REGION Network 68: Alarm - Under Range
   RUNG wire#powerrail
      Contact( #Timers.UR_HLD.Q )
      S_SR(operand := #HMI.Alarm.Alarms.%X7, r1 := wire#w1)
   END_RUNG
   RUNG wire#powerrail
      I_Contact( #Timers.UR_HLD.Q )
      { S7_Templates := "SrcType := Real"; S7_GenerateENO := "TRUE" } Add(in1 := #Admin.SCL.UR, in2 := #Retain.HMI.Config.SP.HYS.UR, out => #Admin.HYS.UR)
      { S7_Templates := "SrcType := Real" } GE_Contact(in1 := #RAIVR_1_1, in2 := #Admin.HYS.UR)
   END_RUNG wire#w1
   RUNG wire#powerrail
      I_Contact( #Retain.HMI.Config.Alarms.%X7 )
   END_RUNG wire#w1
   // the same network as SCL:
   // ENO of a box is taken as its EN; it also drops when the box reports an error
   IF NOT #Timers.UR_HLD.Q THEN #Admin.HYS.UR := #Admin.SCL.UR + #Retain.HMI.Config.SP.HYS.UR; END_IF;
   IF #Timers.UR_HLD.Q THEN
       #HMI.Alarm.Alarms.%X7 := TRUE;   // SR flip-flop
   END_IF;
   IF (NOT #Timers.UR_HLD.Q AND (#RAIVR_1_1 >= #Admin.HYS.UR)) OR NOT #Retain.HMI.Config.Alarms.%X7 THEN
       #HMI.Alarm.Alarms.%X7 := FALSE;
   END_IF;
END_REGION

REGION Network 69: Alarm - Fault
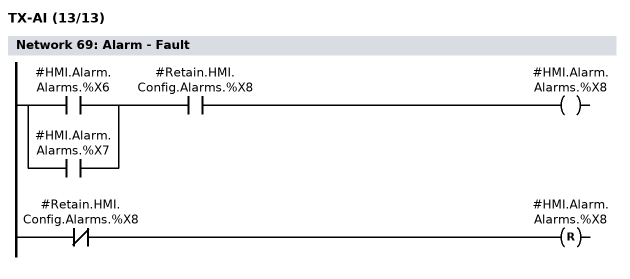
   RUNG wire#powerrail
      Contact( #HMI.Alarm.Alarms.%X6 )
      wire#w1
      Contact( #Retain.HMI.Config.Alarms.%X8 )
      Coil( #HMI.Alarm.Alarms.%X8 )
   END_RUNG
   RUNG wire#powerrail
      Contact( #HMI.Alarm.Alarms.%X7 )
   END_RUNG wire#w1
   RUNG wire#powerrail
      I_Contact( #Retain.HMI.Config.Alarms.%X8 )
      R_Coil( #HMI.Alarm.Alarms.%X8 )
   END_RUNG
   // the same network as SCL:
   #HMI.Alarm.Alarms.%X8 := (#HMI.Alarm.Alarms.%X6 OR #HMI.Alarm.Alarms.%X7) AND #Retain.HMI.Config.Alarms.%X8;
   IF NOT #Retain.HMI.Config.Alarms.%X8 THEN #HMI.Alarm.Alarms.%X8 := FALSE; END_IF;
END_REGION

REGION Network 70 (SCL)
   #Alarms.HighHighHigh := #HMI.Alarm.Alarms.%X0;
   #Alarms.HighHigh := #HMI.Alarm.Alarms.%X1;
   #Alarms.High := #HMI.Alarm.Alarms.%X2;
   #Alarms.Low := #HMI.Alarm.Alarms.%X3;
   #Alarms.LowLow := #HMI.Alarm.Alarms.%X4;
   //#HMI.Alarm.Alarms.%X4:=#Alarms.LowLow;
   #Alarms.LowLowLow := #HMI.Alarm.Alarms.%X5;
   #Alarms.OverRange := #HMI.Alarm.Alarms.%X6;
   #Alarms.UnderRange := #HMI.Alarm.Alarms.%X7;
   #Alarms.TransmitterFault := #HMI.Alarm.Alarms.%X8;
END_REGION
END_FUNCTION_BLOCK

FUNCTION_BLOCK "TX-AI_Basic"   // FB805, LAD
TITLE = SSAC Basic Analog Trasmitter Function Block
{ S7_Optimized_Access := 'FALSE' }
VERSION : 1.0
// Default mode 0 starts at  network 4
   VAR_INPUT
      Mode : Int;   // TX Mode - 0 = 4-20 mA / 1 = Int Math (RTD/TC) / 2 = Real Input Conversion
      RAIVI : Int;   // Raw Analog Input Value INT
      RAIVR : Real;   // Raw Analog Input Value REAL
   END_VAR
   VAR_OUTPUT
      SAI : Real;   // Compensated Scaled Analog Value
   END_VAR
   VAR
      HMI : Struct   // Alarms
         Status : Struct
            USAV : Real;   // Uncompensated Scaled Analog Value
            NV : Real;   // Normalized Value
         END_STRUCT;
         Alarm : Struct
            Alarms : Word;
         END_STRUCT;
         Diag : Struct   // Diagnostics
            SV : Real;   // Simulation Value
         END_STRUCT;
      END_STRUCT;
      Retain : Struct
         HMI : Struct
            Config : Struct   // Settings
               RIMXV : Real := 27648.0;   // Raw Input Maximum Value (Used for Sqrt)
               RIMNV : Real;   // Raw Input Minimum Value (Used for Sqrt)
               ESMXV : Real := 100.0;   // Engineering/Scaled Maximum Value
               ESMNV : Real;   // Engineering/Scaled Minimum Value
               SAM : Bool;   // Substitution Activation Mode
               SAV : Real := -999999.0;   // Substitution Value during a limit input value trip
               SP : Struct   // Setpoints
                  Limits : Struct
                     HHH : Real := 95.0;   // HHH Limit Setpoint
                     HH : Real := 90.0;   // HH Limit Setpoint
                     H : Real := 80.0;   // HH Limit Setpoint
                     L : Real := 20.0;   // L Limit Setpoint
                     LL : Real := 10.0;   // LL Limit Setpoint
                     LLL : Real := 5.0;   // LLL Limit Setpoint
                     "OR" : Real := 5.0;   // Over range value
                     UR : Real := 5.0;   // Under range value
                  END_STRUCT;
                  HYS : Struct   // Hysteresis
                     Global : Real;   // Hysteresis global value, only valid when greater than or equal to 0
                     HHH : Real := 1.0;   // Hysteresis Setpoint - High High High
                     HH : Real := 1.0;   // Hysteresis Setpoint - High High
                     H : Real := 1.0;   // Hysteresis Setpoint - High
                     L : Real := 1.0;   // Hysteresis Setpoint - Low
                     LL : Real := 1.0;   // Hysteresis Setpoint - Low Low
                     LLL : Real := 1.0;   // Hysteresis Setpoint - Low Low Low
                     "OR" : Real := 1.0;   // Hysteresis Setpoint - Over Range
                     UR : Real := 1.0;   // Hysteresis Setpoint - Under Range
                  END_STRUCT;
                  SUB_ON : Bool;   // Substitution Activation
               END_STRUCT;
               PT : Struct   // Setpoints
                  HLD : Struct   // Hold
                     Global : Time;   // Hold PT global value, only valid when not equal to 0
                     AHHH : Time := t#5s;   // Alarm Debounce
                     AHH : Time := t#5s;   // Alarm Debounce
                     AH : Time := t#5s;   // Alarm Debounce
                     AL : Time := t#5s;   // Alarm Debounce
                     ALL : Time := t#5s;   // Alarm Debounce
                     ALLL : Time := t#5s;   // Alarm Debounce
                     "OR" : Time := t#5s;   // Over range hold
                     UR : Time := t#5s;   // Under range hold
                  END_STRUCT;
                  DBNC : Struct   // Debounce
                     Global : Time;   // Debounce PT global value, only valid when not equal to 0
                     AHHH : Time := t#5s;   // Alarm Debounce
                     AHH : Time := t#5s;   // Alarm Debounce
                     AH : Time := t#5s;   // Alarm Debounce
                     AL : Time := t#5s;   // Alarm Debounce
                     ALL : Time := t#5s;   // Alarm Debounce
                     ALLL : Time := t#5s;   // Alarm Debounce
                     "OR" : Time := t#5s;   // Over range debounce
                     UR : Time := t#5s;   // Under range debounce
                  END_STRUCT;
               END_STRUCT;
               Alarms : Word := 16#03DE;
            END_STRUCT;
         END_STRUCT;
      END_STRUCT;
      Admin : Struct   // Admin configurations
         SCL : Struct   // Scale Values
            RDP : Real := 10.0;   // RTD Decimal Places
            RRIMD : Real := 1.0;   // Raw Real input Math divider
            "OR" : Real;   // Over Range Value
            UR : Real;   // Under Range Value
            SAIV : Real;   // Scaled Analog Input Value
         END_STRUCT;
         HYS : Struct   // Hysteresis - Computed Values
            "OR" : Real;   // Hysteresis Value - Over Range
            UR : Real;   // Hysteresis Value - Under Range
         END_STRUCT;
      END_STRUCT;
      Alarms : Struct
         HighHighHigh : Bool;
         HighHigh : Bool;
         High : Bool;
         Low : Bool;
         LowLow : Bool;
         LowLowLow : Bool;
         TransmitterFault : Bool;
         UnderRange : Bool;
         OverRange : Bool;
      END_STRUCT;
      Timers : Struct
         OR_DB : TON_TIME;   // Over Range Debounce
         UR_DB : TON_TIME;   // Under Range DB
         OR_HLD : TOF_TIME;   // Over Range Hold
         UR_HLD : TOF_TIME;   // Under Range Hold
         DBNC : Struct
            HHH : TON_TIME;
            HH : TON_TIME;
            H : TON_TIME;
            L : TON_TIME;
            LL : TON_TIME;
            LLL : TON_TIME;
         END_STRUCT;
         HOLD : Struct
            HHH : TOF_TIME;
            HH : TOF_TIME;
            H : TOF_TIME;
            L : TOF_TIME;
            LL : TOF_TIME;
            LLL : TOF_TIME;
         END_STRUCT;
      END_STRUCT;
   END_VAR
   VAR_TEMP
      SRV : Real;
      RAIDI : DInt;   // Raw Analog Input DINT
      RAIR : Real;   // Raw Analog Input REAL
      RAIVR_1 : DInt;
      RAIVR_1_1 : Real;
      ValuePerPoint : Real;
      ValueAddRaw : Real;
      voidTime : Word;
   END_VAR
   VAR_TEMP   // added for the SCL form of the ladder/FBD networks
      _w1 : Bool;
   END_VAR
BEGIN

REGION Network 1: Transmitter Mode 1 = Int Math or RTD
   // MD1 Jump to network 7
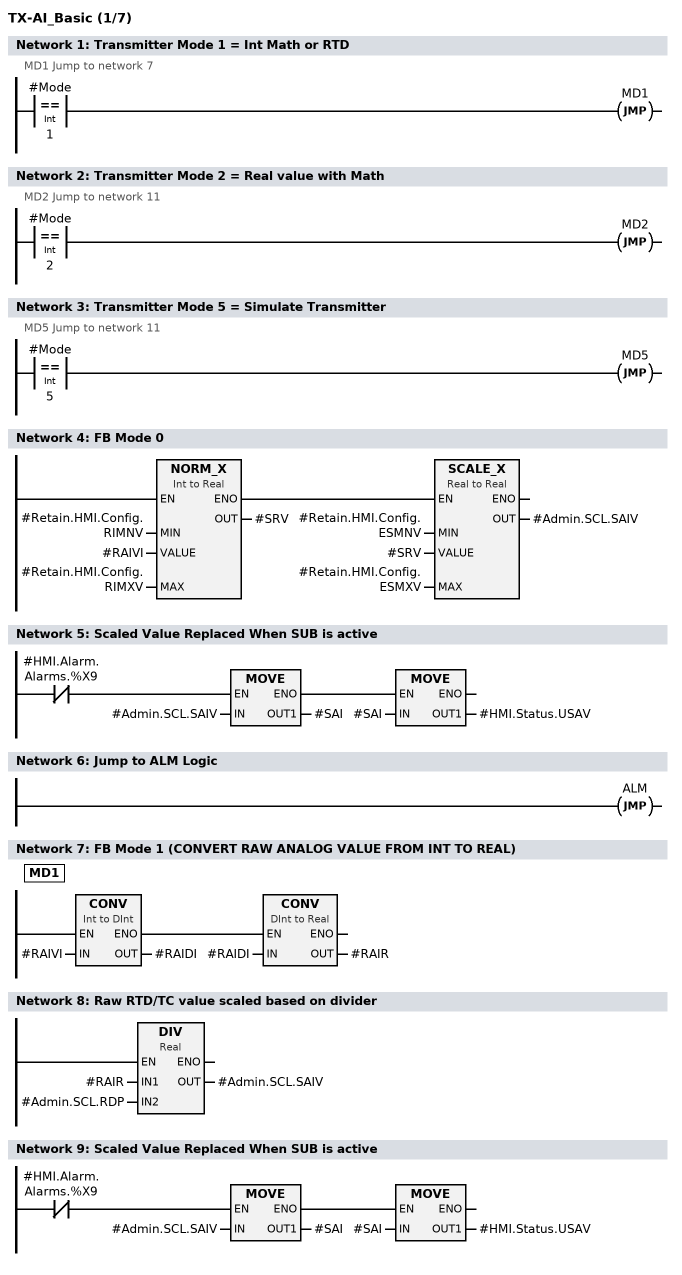
   RUNG wire#powerrail
      { S7_Templates := "SrcType := Int" } EQ_Contact(in1 := #Mode, in2 := 1)
      JumpCoil( MD1 )
   END_RUNG
   // the same network as SCL:
   IF #Mode = 1 THEN GOTO MD1; END_IF;
END_REGION

REGION Network 2: Transmitter Mode 2 = Real value with Math
   // MD2 Jump to network 11
   RUNG wire#powerrail
      { S7_Templates := "SrcType := Int" } EQ_Contact(in1 := #Mode, in2 := 2)
      JumpCoil( MD2 )
   END_RUNG
   // the same network as SCL:
   IF #Mode = 2 THEN GOTO MD2; END_IF;
END_REGION

REGION Network 3: Transmitter Mode 5 = Simulate Transmitter
   // MD5 Jump to network 11
   RUNG wire#powerrail
      { S7_Templates := "SrcType := Int" } EQ_Contact(in1 := #Mode, in2 := 5)
      JumpCoil( MD5 )
   END_RUNG
   // the same network as SCL:
   IF #Mode = 5 THEN GOTO MD5; END_IF;
END_REGION

REGION Network 4: FB Mode 0
   RUNG wire#powerrail
      { S7_Templates := "[SrcType := Int, DestType := Real]" } Normalize(min := #Retain.HMI.Config.RIMNV, value := #RAIVI, max := #Retain.HMI.Config.RIMXV, out => #SRV)
      { S7_Templates := "[SrcType := Real, DestType := Real]" } Scale(min := #Retain.HMI.Config.ESMNV, value := #SRV, max := #Retain.HMI.Config.ESMXV, out => #Admin.SCL.SAIV)
   END_RUNG
   // the same network as SCL:
   #SRV := NORM_X(MIN := #Retain.HMI.Config.RIMNV, VALUE := #RAIVI, MAX := #Retain.HMI.Config.RIMXV);
   #Admin.SCL.SAIV := SCALE_X(MIN := #Retain.HMI.Config.ESMNV, VALUE := #SRV, MAX := #Retain.HMI.Config.ESMXV);
END_REGION

REGION Network 5: Scaled Value Replaced When SUB is active
   RUNG wire#powerrail
      I_Contact( #HMI.Alarm.Alarms.%X9 )
      { S7_GenerateENO := "TRUE" } Move(in := #Admin.SCL.SAIV, out1 => #SAI)
      { S7_GenerateENO := "TRUE" } Move(in := #SAI, out1 => #HMI.Status.USAV)
   END_RUNG
   // the same network as SCL:
   // ENO of a box is taken as its EN; it also drops when the box reports an error
   IF NOT #HMI.Alarm.Alarms.%X9 THEN
       #SAI := #Admin.SCL.SAIV;
       #HMI.Status.USAV := #SAI;
   END_IF;
END_REGION

REGION Network 6: Jump to ALM Logic
   RUNG wire#powerrail
      JumpCoil( ALM )
   END_RUNG
   // the same network as SCL:
   GOTO ALM;
END_REGION

REGION Network 7: FB Mode 1 (CONVERT RAW ANALOG VALUE FROM INT TO REAL)
   Label( MD1 )
   RUNG wire#powerrail
      { S7_Templates := "[SrcType := Int, DestType := DInt]"; S7_GenerateENO := "TRUE" } Convert(in := #RAIVI, out => #RAIDI)
      { S7_Templates := "[SrcType := DInt, DestType := Real]"; S7_GenerateENO := "TRUE" } Convert(in := #RAIDI, out => #RAIR)
   END_RUNG
   // the same network as SCL:
   // ENO of a box is taken as its EN; it also drops when the box reports an error
   MD1:
   #RAIDI := INT_TO_DINT(#RAIVI);
   #RAIR := DINT_TO_REAL(#RAIDI);
END_REGION

REGION Network 8: Raw RTD/TC value scaled based on divider
   RUNG wire#powerrail
      { S7_Templates := "SrcType := Real"; S7_GenerateENO := "TRUE" } Div(in1 := #RAIR, in2 := #Admin.SCL.RDP, out => #Admin.SCL.SAIV)
   END_RUNG
   // the same network as SCL:
   #Admin.SCL.SAIV := #RAIR / #Admin.SCL.RDP;
END_REGION

REGION Network 9: Scaled Value Replaced When SUB is active
   RUNG wire#powerrail
      I_Contact( #HMI.Alarm.Alarms.%X9 )
      { S7_GenerateENO := "TRUE" } Move(in := #Admin.SCL.SAIV, out1 => #SAI)
      Move(in := #SAI, out1 => #HMI.Status.USAV)
   END_RUNG
   // the same network as SCL:
   // ENO of a box is taken as its EN; it also drops when the box reports an error
   IF NOT #HMI.Alarm.Alarms.%X9 THEN
       #SAI := #Admin.SCL.SAIV;
       #HMI.Status.USAV := #SAI;
   END_IF;
END_REGION

REGION Network 10: Jump to ALM Logic
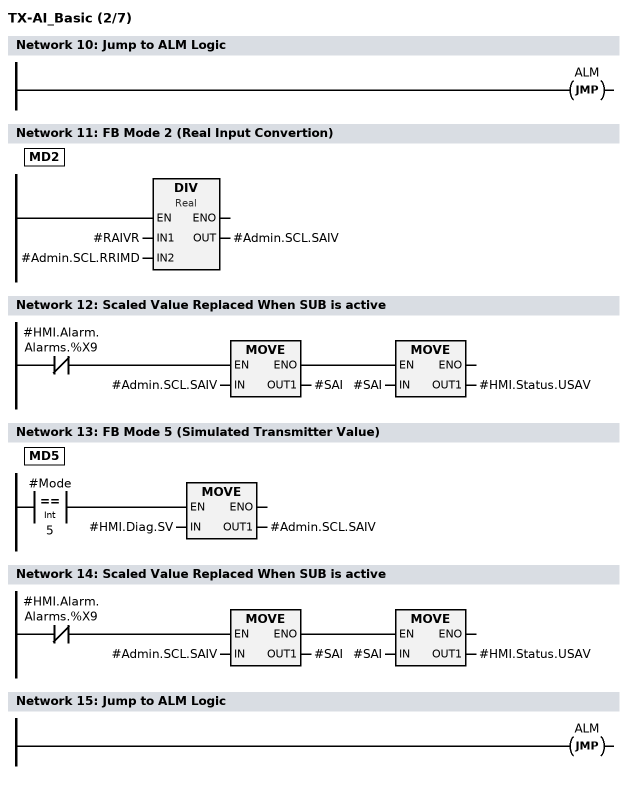
   RUNG wire#powerrail
      JumpCoil( ALM )
   END_RUNG
   // the same network as SCL:
   GOTO ALM;
END_REGION

REGION Network 11: FB Mode 2 (Real Input Convertion)
   Label( MD2 )
   RUNG wire#powerrail
      { S7_Templates := "SrcType := Real"; S7_GenerateENO := "TRUE" } Div(in1 := #RAIVR, in2 := #Admin.SCL.RRIMD, out => #Admin.SCL.SAIV)
   END_RUNG
   // the same network as SCL:
   MD2:
   #Admin.SCL.SAIV := #RAIVR / #Admin.SCL.RRIMD;
END_REGION

REGION Network 12: Scaled Value Replaced When SUB is active
   RUNG wire#powerrail
      I_Contact( #HMI.Alarm.Alarms.%X9 )
      { S7_GenerateENO := "TRUE" } Move(in := #Admin.SCL.SAIV, out1 => #SAI)
      Move(in := #SAI, out1 => #HMI.Status.USAV)
   END_RUNG
   // the same network as SCL:
   // ENO of a box is taken as its EN; it also drops when the box reports an error
   IF NOT #HMI.Alarm.Alarms.%X9 THEN
       #SAI := #Admin.SCL.SAIV;
       #HMI.Status.USAV := #SAI;
   END_IF;
END_REGION

REGION Network 13: FB Mode 5 (Simulated Transmitter Value)
   Label( MD5 )
   RUNG wire#powerrail
      { S7_Templates := "SrcType := Int" } EQ_Contact(in1 := #Mode, in2 := 5)
      { S7_GenerateENO := "TRUE" } Move(in := #HMI.Diag.SV, out1 => #Admin.SCL.SAIV)
   END_RUNG
   // the same network as SCL:
   MD5:
   IF #Mode = 5 THEN #Admin.SCL.SAIV := #HMI.Diag.SV; END_IF;
END_REGION

REGION Network 14: Scaled Value Replaced When SUB is active
   RUNG wire#powerrail
      I_Contact( #HMI.Alarm.Alarms.%X9 )
      { S7_GenerateENO := "TRUE" } Move(in := #Admin.SCL.SAIV, out1 => #SAI)
      { S7_GenerateENO := "TRUE" } Move(in := #SAI, out1 => #HMI.Status.USAV)
   END_RUNG
   // the same network as SCL:
   // ENO of a box is taken as its EN; it also drops when the box reports an error
   IF NOT #HMI.Alarm.Alarms.%X9 THEN
       #SAI := #Admin.SCL.SAIV;
       #HMI.Status.USAV := #SAI;
   END_IF;
END_REGION

REGION Network 15: Jump to ALM Logic
   RUNG wire#powerrail
      JumpCoil( ALM )
   END_RUNG
   // the same network as SCL:
   GOTO ALM;
END_REGION

REGION Network 16: Global Hysteresis Setpoint Condition
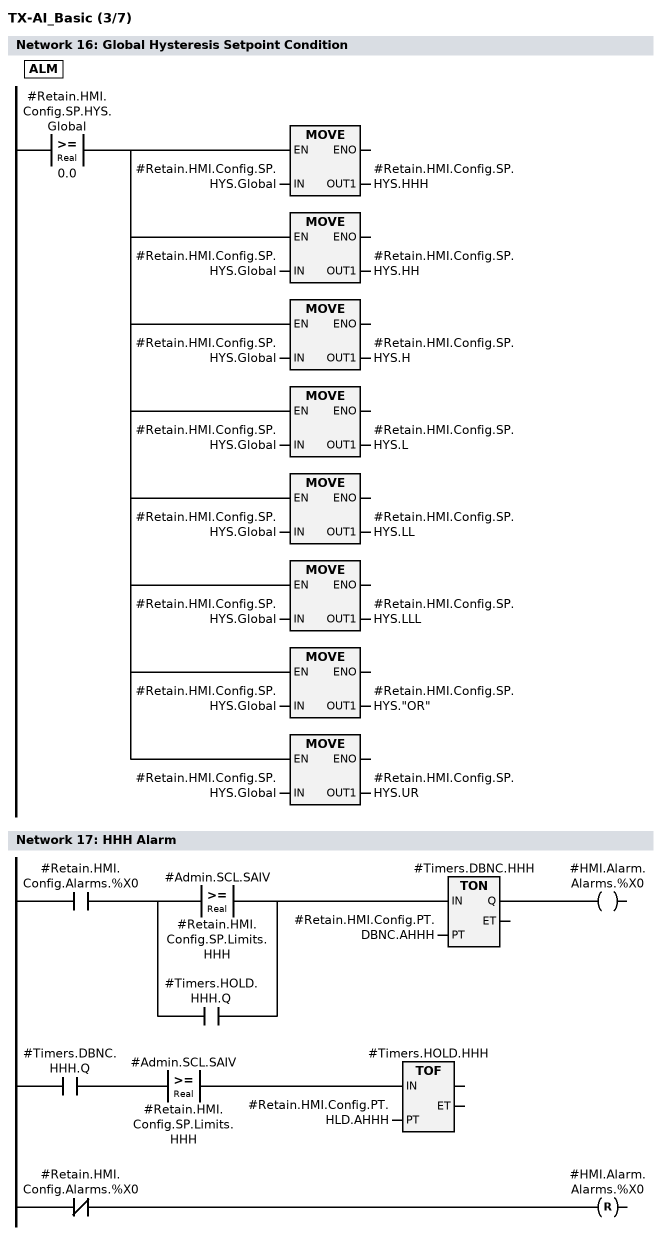
   Label( ALM )
   RUNG wire#powerrail
      { S7_Templates := "SrcType := Real" } GE_Contact(in1 := #Retain.HMI.Config.SP.HYS.Global, in2 := 0.0)
      wire#w1
      { S7_GenerateENO := "TRUE" } Move(in := #Retain.HMI.Config.SP.HYS.Global, out1 => #Retain.HMI.Config.SP.HYS.HHH)
   END_RUNG
   RUNG wire#w1
      { S7_GenerateENO := "TRUE" } Move(in := #Retain.HMI.Config.SP.HYS.Global, out1 => #Retain.HMI.Config.SP.HYS.HH)
   END_RUNG
   RUNG wire#w1
      { S7_GenerateENO := "TRUE" } Move(in := #Retain.HMI.Config.SP.HYS.Global, out1 => #Retain.HMI.Config.SP.HYS.H)
   END_RUNG
   RUNG wire#w1
      { S7_GenerateENO := "TRUE" } Move(in := #Retain.HMI.Config.SP.HYS.Global, out1 => #Retain.HMI.Config.SP.HYS.L)
   END_RUNG
   RUNG wire#w1
      { S7_GenerateENO := "TRUE" } Move(in := #Retain.HMI.Config.SP.HYS.Global, out1 => #Retain.HMI.Config.SP.HYS.LL)
   END_RUNG
   RUNG wire#w1
      { S7_GenerateENO := "TRUE" } Move(in := #Retain.HMI.Config.SP.HYS.Global, out1 => #Retain.HMI.Config.SP.HYS.LLL)
   END_RUNG
   RUNG wire#w1
      { S7_GenerateENO := "TRUE" } Move(in := #Retain.HMI.Config.SP.HYS.Global, out1 => #Retain.HMI.Config.SP.HYS."OR")
   END_RUNG
   RUNG wire#w1
      { S7_GenerateENO := "TRUE" } Move(in := #Retain.HMI.Config.SP.HYS.Global, out1 => #Retain.HMI.Config.SP.HYS.UR)
   END_RUNG
   // the same network as SCL:
   ALM:
   IF #Retain.HMI.Config.SP.HYS.Global >= 0.0 THEN
       #Retain.HMI.Config.SP.HYS.HHH := #Retain.HMI.Config.SP.HYS.Global;
       #Retain.HMI.Config.SP.HYS.HH := #Retain.HMI.Config.SP.HYS.Global;
       #Retain.HMI.Config.SP.HYS.H := #Retain.HMI.Config.SP.HYS.Global;
       #Retain.HMI.Config.SP.HYS.L := #Retain.HMI.Config.SP.HYS.Global;
       #Retain.HMI.Config.SP.HYS.LL := #Retain.HMI.Config.SP.HYS.Global;
       #Retain.HMI.Config.SP.HYS.LLL := #Retain.HMI.Config.SP.HYS.Global;
       #Retain.HMI.Config.SP.HYS."OR" := #Retain.HMI.Config.SP.HYS.Global;
       #Retain.HMI.Config.SP.HYS.UR := #Retain.HMI.Config.SP.HYS.Global;
   END_IF;
END_REGION

REGION Network 17: HHH Alarm
   #Timers.DBNC.HHH.TON(IN := #Retain.HMI.Config.Alarms.%X0 AND ((#Admin.SCL.SAIV >= #Retain.HMI.Config.SP.Limits.HHH) OR #Timers.HOLD.HHH.Q),
                        PT := #Retain.HMI.Config.PT.DBNC.AHHH);
   #HMI.Alarm.Alarms.%X0 := #Timers.DBNC.HHH.Q;
   #Timers.HOLD.HHH.TOF(IN := #Timers.DBNC.HHH.Q AND (#Admin.SCL.SAIV >= #Retain.HMI.Config.SP.Limits.HHH),
                        PT := #Retain.HMI.Config.PT.HLD.AHHH);
   IF NOT #Retain.HMI.Config.Alarms.%X0 THEN #HMI.Alarm.Alarms.%X0 := FALSE; END_IF;
END_REGION

REGION Network 18: HH Alarm
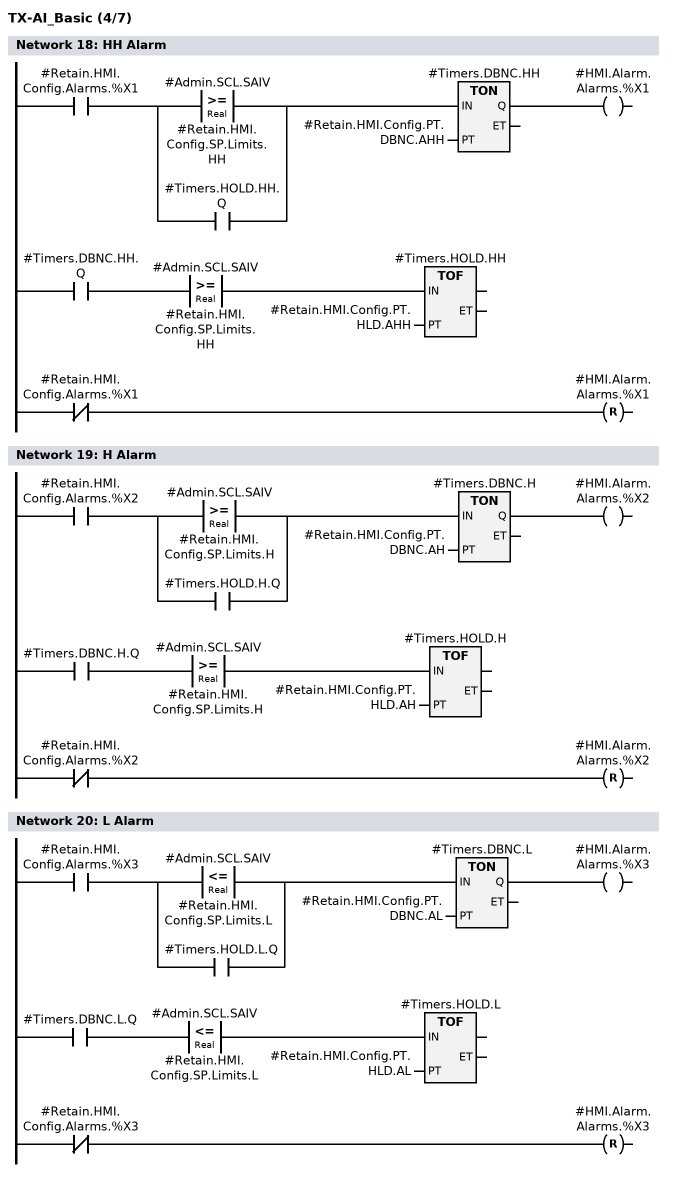
   #Timers.DBNC.HH.TON(IN := #Retain.HMI.Config.Alarms.%X1 AND ((#Admin.SCL.SAIV >= #Retain.HMI.Config.SP.Limits.HH) OR #Timers.HOLD.HH.Q),
                       PT := #Retain.HMI.Config.PT.DBNC.AHH);
   #HMI.Alarm.Alarms.%X1 := #Timers.DBNC.HH.Q;
   #Timers.HOLD.HH.TOF(IN := #Timers.DBNC.HH.Q AND (#Admin.SCL.SAIV >= #Retain.HMI.Config.SP.Limits.HH),
                       PT := #Retain.HMI.Config.PT.HLD.AHH);
   IF NOT #Retain.HMI.Config.Alarms.%X1 THEN #HMI.Alarm.Alarms.%X1 := FALSE; END_IF;
END_REGION

REGION Network 19: H Alarm
   #Timers.DBNC.H.TON(IN := #Retain.HMI.Config.Alarms.%X2 AND ((#Admin.SCL.SAIV >= #Retain.HMI.Config.SP.Limits.H) OR #Timers.HOLD.H.Q),
                      PT := #Retain.HMI.Config.PT.DBNC.AH);
   #HMI.Alarm.Alarms.%X2 := #Timers.DBNC.H.Q;
   #Timers.HOLD.H.TOF(IN := #Timers.DBNC.H.Q AND (#Admin.SCL.SAIV >= #Retain.HMI.Config.SP.Limits.H),
                      PT := #Retain.HMI.Config.PT.HLD.AH);
   IF NOT #Retain.HMI.Config.Alarms.%X2 THEN #HMI.Alarm.Alarms.%X2 := FALSE; END_IF;
END_REGION

REGION Network 20: L Alarm
   #Timers.DBNC.L.TON(IN := #Retain.HMI.Config.Alarms.%X3 AND ((#Admin.SCL.SAIV <= #Retain.HMI.Config.SP.Limits.L) OR #Timers.HOLD.L.Q),
                      PT := #Retain.HMI.Config.PT.DBNC.AL);
   #HMI.Alarm.Alarms.%X3 := #Timers.DBNC.L.Q;
   #Timers.HOLD.L.TOF(IN := #Timers.DBNC.L.Q AND (#Admin.SCL.SAIV <= #Retain.HMI.Config.SP.Limits.L),
                      PT := #Retain.HMI.Config.PT.HLD.AL);
   IF NOT #Retain.HMI.Config.Alarms.%X3 THEN #HMI.Alarm.Alarms.%X3 := FALSE; END_IF;
END_REGION

REGION Network 21: LL Alarm
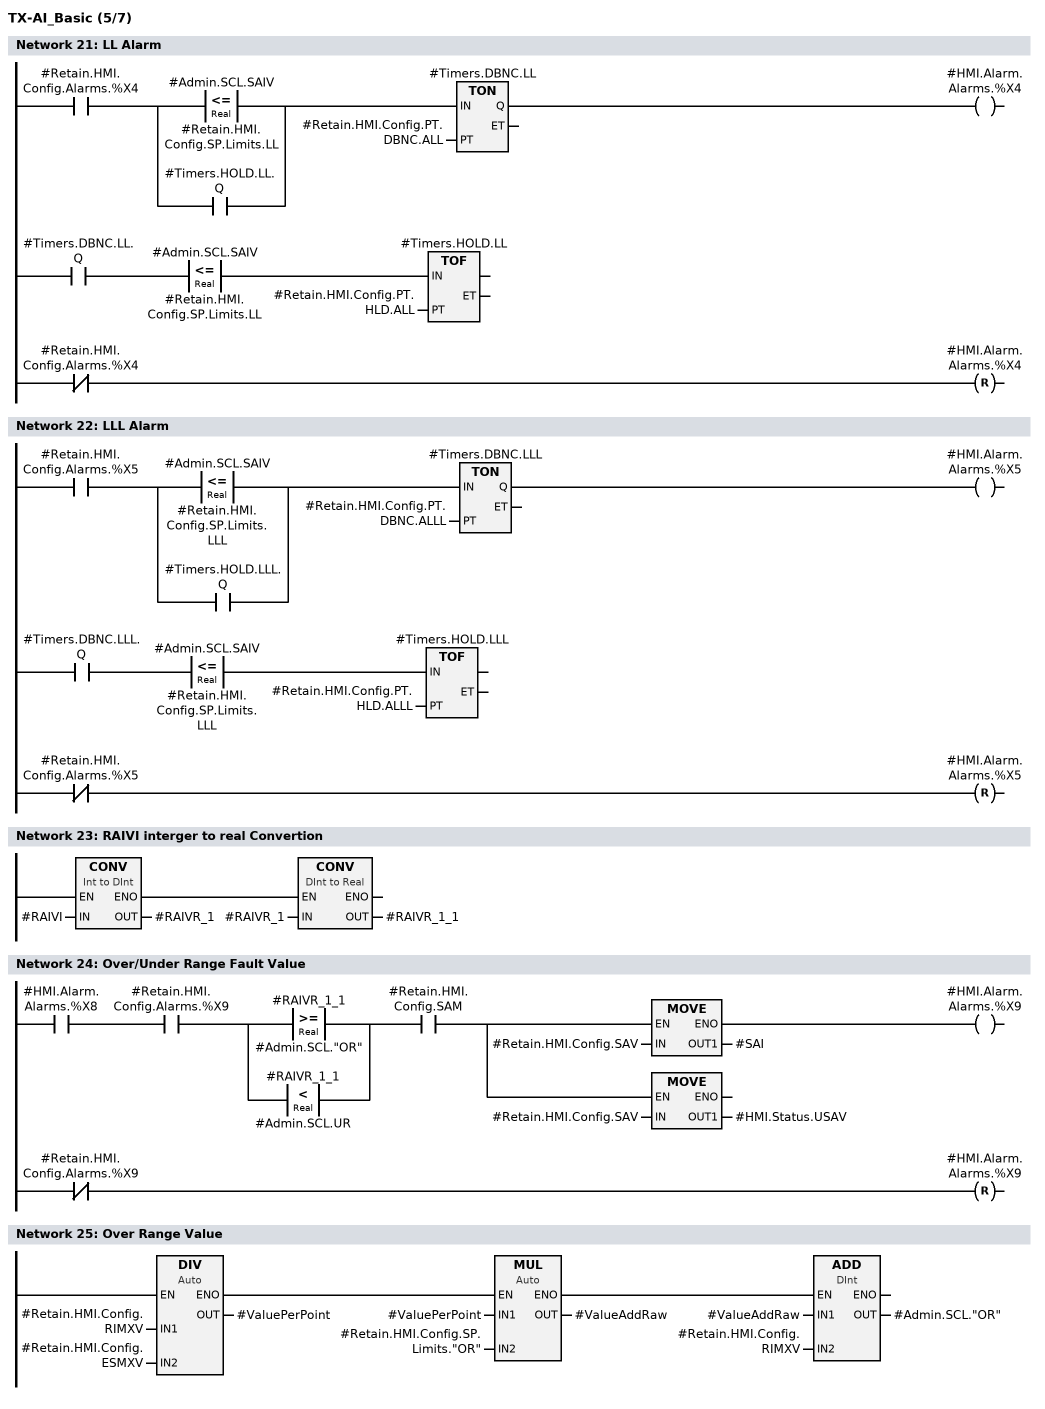
   #Timers.DBNC.LL.TON(IN := #Retain.HMI.Config.Alarms.%X4 AND ((#Admin.SCL.SAIV <= #Retain.HMI.Config.SP.Limits.LL) OR #Timers.HOLD.LL.Q),
                       PT := #Retain.HMI.Config.PT.DBNC.ALL);
   #HMI.Alarm.Alarms.%X4 := #Timers.DBNC.LL.Q;
   #Timers.HOLD.LL.TOF(IN := #Timers.DBNC.LL.Q AND (#Admin.SCL.SAIV <= #Retain.HMI.Config.SP.Limits.LL),
                       PT := #Retain.HMI.Config.PT.HLD.ALL);
   IF NOT #Retain.HMI.Config.Alarms.%X4 THEN #HMI.Alarm.Alarms.%X4 := FALSE; END_IF;
END_REGION

REGION Network 22: LLL Alarm
   #Timers.DBNC.LLL.TON(IN := #Retain.HMI.Config.Alarms.%X5 AND ((#Admin.SCL.SAIV <= #Retain.HMI.Config.SP.Limits.LLL) OR #Timers.HOLD.LLL.Q),
                        PT := #Retain.HMI.Config.PT.DBNC.ALLL);
   #HMI.Alarm.Alarms.%X5 := #Timers.DBNC.LLL.Q;
   #Timers.HOLD.LLL.TOF(IN := #Timers.DBNC.LLL.Q AND (#Admin.SCL.SAIV <= #Retain.HMI.Config.SP.Limits.LLL),
                        PT := #Retain.HMI.Config.PT.HLD.ALLL);
   IF NOT #Retain.HMI.Config.Alarms.%X5 THEN #HMI.Alarm.Alarms.%X5 := FALSE; END_IF;
END_REGION

REGION Network 23: RAIVI interger to real Convertion
   RUNG wire#powerrail
      { S7_Templates := "[SrcType := Int, DestType := DInt]"; S7_GenerateENO := "TRUE" } Convert(in := #RAIVI, out => #RAIVR_1)
      { S7_Templates := "[SrcType := DInt, DestType := Real]"; S7_GenerateENO := "TRUE" } Convert(in := #RAIVR_1, out => #RAIVR_1_1)
   END_RUNG
   // the same network as SCL:
   // ENO of a box is taken as its EN; it also drops when the box reports an error
   #RAIVR_1 := INT_TO_DINT(#RAIVI);
   #RAIVR_1_1 := DINT_TO_REAL(#RAIVR_1);
END_REGION

REGION Network 24: Over/Under Range Fault Value
   RUNG wire#powerrail
      Contact( #HMI.Alarm.Alarms.%X8 )
      Contact( #Retain.HMI.Config.Alarms.%X9 )
      wire#w1
      { S7_Templates := "SrcType := Real" } GE_Contact(in1 := #RAIVR_1_1, in2 := #Admin.SCL."OR")
      wire#w2
      Contact( #Retain.HMI.Config.SAM )
      wire#w3
      { S7_GenerateENO := "TRUE" } Move(in := #Retain.HMI.Config.SAV, out1 => #SAI)
      Coil( #HMI.Alarm.Alarms.%X9 )
   END_RUNG
   RUNG wire#w1
      { S7_Templates := "SrcType := Real" } LT_Contact(in1 := #RAIVR_1_1, in2 := #Admin.SCL.UR)
   END_RUNG wire#w2
   RUNG wire#w3
      { S7_GenerateENO := "TRUE" } Move(in := #Retain.HMI.Config.SAV, out1 => #HMI.Status.USAV)
   END_RUNG
   RUNG wire#powerrail
      I_Contact( #Retain.HMI.Config.Alarms.%X9 )
      R_Coil( #HMI.Alarm.Alarms.%X9 )
   END_RUNG
   // the same network as SCL:
   // ENO of a box is taken as its EN; it also drops when the box reports an error
   #_w1 := #HMI.Alarm.Alarms.%X8 AND #Retain.HMI.Config.Alarms.%X9 AND ((#RAIVR_1_1 >= #Admin.SCL."OR") OR (#RAIVR_1_1 < #Admin.SCL.UR)) AND #Retain.HMI.Config.SAM;
   IF #_w1 THEN #SAI := #Retain.HMI.Config.SAV; END_IF;
   #HMI.Alarm.Alarms.%X9 := #_w1;
   IF #_w1 THEN #HMI.Status.USAV := #Retain.HMI.Config.SAV; END_IF;
   IF NOT #Retain.HMI.Config.Alarms.%X9 THEN #HMI.Alarm.Alarms.%X9 := FALSE; END_IF;
END_REGION

REGION Network 25: Over Range Value
   RUNG wire#powerrail
      Div(in1 := #Retain.HMI.Config.RIMXV, in2 := #Retain.HMI.Config.ESMXV, out => #ValuePerPoint)
      Mul(in1 := #ValuePerPoint, in2 := #Retain.HMI.Config.SP.Limits."OR", out => #ValueAddRaw)
      { S7_Templates := "SrcType := DInt"; S7_GenerateENO := "TRUE" } Add(in1 := #ValueAddRaw, in2 := #Retain.HMI.Config.RIMXV, out => #Admin.SCL."OR")
   END_RUNG
   // the same network as SCL:
   #ValuePerPoint := #Retain.HMI.Config.RIMXV / #Retain.HMI.Config.ESMXV;
   #ValueAddRaw := #ValuePerPoint * #Retain.HMI.Config.SP.Limits."OR";
   #Admin.SCL."OR" := #ValueAddRaw + #Retain.HMI.Config.RIMXV;
END_REGION

REGION Network 26: Under Range Value
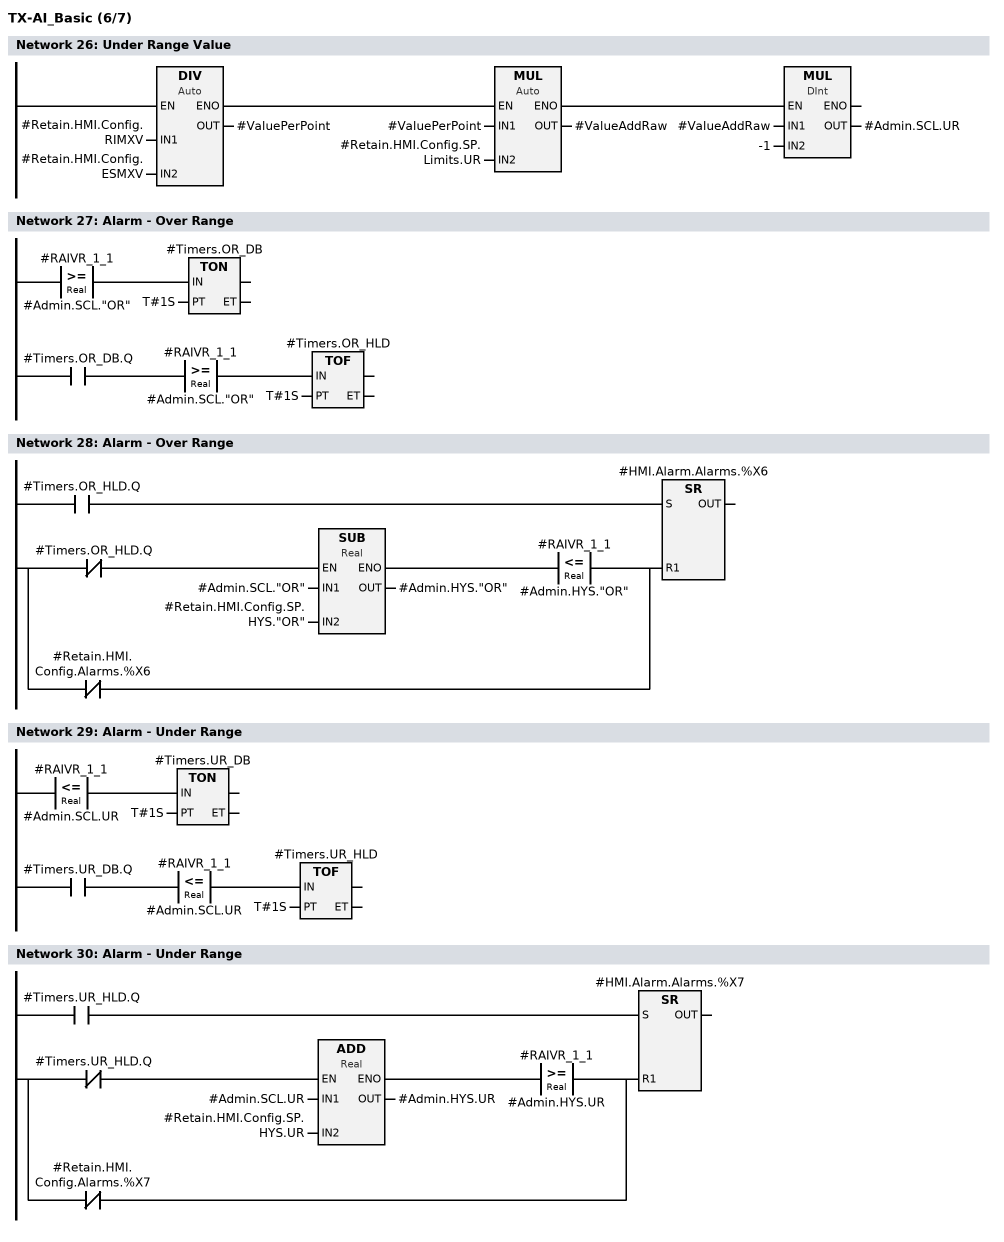
   RUNG wire#powerrail
      Div(in1 := #Retain.HMI.Config.RIMXV, in2 := #Retain.HMI.Config.ESMXV, out => #ValuePerPoint)
      Mul(in1 := #ValuePerPoint, in2 := #Retain.HMI.Config.SP.Limits.UR, out => #ValueAddRaw)
      { S7_Templates := "SrcType := DInt"; S7_GenerateENO := "TRUE" } Mul(in1 := #ValueAddRaw, in2 := -1, out => #Admin.SCL.UR)
   END_RUNG
   // the same network as SCL:
   #ValuePerPoint := #Retain.HMI.Config.RIMXV / #Retain.HMI.Config.ESMXV;
   #ValueAddRaw := #ValuePerPoint * #Retain.HMI.Config.SP.Limits.UR;
   #Admin.SCL.UR := #ValueAddRaw * (-1);
END_REGION

REGION Network 27: Alarm - Over Range
   #Timers.OR_DB.TON(IN := #RAIVR_1_1 >= #Admin.SCL."OR", PT := T#1S);
   #Timers.OR_HLD.TOF(IN := #Timers.OR_DB.Q AND (#RAIVR_1_1 >= #Admin.SCL."OR"), PT := T#1S);
END_REGION

REGION Network 28: Alarm - Over Range
   RUNG wire#powerrail
      Contact( #Timers.OR_HLD.Q )
      S_SR(operand := #HMI.Alarm.Alarms.%X6, r1 := wire#w1)
   END_RUNG
   RUNG wire#powerrail
      I_Contact( #Timers.OR_HLD.Q )
      { S7_Templates := "SrcType := Real"; S7_GenerateENO := "TRUE" } Sub(in1 := #Admin.SCL."OR", in2 := #Retain.HMI.Config.SP.HYS."OR", out => #Admin.HYS."OR")
      { S7_Templates := "SrcType := Real" } LE_Contact(in1 := #RAIVR_1_1, in2 := #Admin.HYS."OR")
   END_RUNG wire#w1
   RUNG wire#powerrail
      I_Contact( #Retain.HMI.Config.Alarms.%X6 )
   END_RUNG wire#w1
   // the same network as SCL:
   // ENO of a box is taken as its EN; it also drops when the box reports an error
   IF NOT #Timers.OR_HLD.Q THEN #Admin.HYS."OR" := #Admin.SCL."OR" - #Retain.HMI.Config.SP.HYS."OR"; END_IF;
   IF #Timers.OR_HLD.Q THEN
       #HMI.Alarm.Alarms.%X6 := TRUE;   // SR flip-flop
   END_IF;
   IF (NOT #Timers.OR_HLD.Q AND (#RAIVR_1_1 <= #Admin.HYS."OR")) OR NOT #Retain.HMI.Config.Alarms.%X6 THEN
       #HMI.Alarm.Alarms.%X6 := FALSE;
   END_IF;
END_REGION

REGION Network 29: Alarm - Under Range
   #Timers.UR_DB.TON(IN := #RAIVR_1_1 <= #Admin.SCL.UR, PT := T#1S);
   #Timers.UR_HLD.TOF(IN := #Timers.UR_DB.Q AND (#RAIVR_1_1 <= #Admin.SCL.UR), PT := T#1S);
END_REGION

REGION Network 30: Alarm - Under Range
   RUNG wire#powerrail
      Contact( #Timers.UR_HLD.Q )
      S_SR(operand := #HMI.Alarm.Alarms.%X7, r1 := wire#w1)
   END_RUNG
   RUNG wire#powerrail
      I_Contact( #Timers.UR_HLD.Q )
      { S7_Templates := "SrcType := Real"; S7_GenerateENO := "TRUE" } Add(in1 := #Admin.SCL.UR, in2 := #Retain.HMI.Config.SP.HYS.UR, out => #Admin.HYS.UR)
      { S7_Templates := "SrcType := Real" } GE_Contact(in1 := #RAIVR_1_1, in2 := #Admin.HYS.UR)
   END_RUNG wire#w1
   RUNG wire#powerrail
      I_Contact( #Retain.HMI.Config.Alarms.%X7 )
   END_RUNG wire#w1
   // the same network as SCL:
   // ENO of a box is taken as its EN; it also drops when the box reports an error
   IF NOT #Timers.UR_HLD.Q THEN #Admin.HYS.UR := #Admin.SCL.UR + #Retain.HMI.Config.SP.HYS.UR; END_IF;
   IF #Timers.UR_HLD.Q THEN
       #HMI.Alarm.Alarms.%X7 := TRUE;   // SR flip-flop
   END_IF;
   IF (NOT #Timers.UR_HLD.Q AND (#RAIVR_1_1 >= #Admin.HYS.UR)) OR NOT #Retain.HMI.Config.Alarms.%X7 THEN
       #HMI.Alarm.Alarms.%X7 := FALSE;
   END_IF;
END_REGION

REGION Network 31: Alarm - Fault
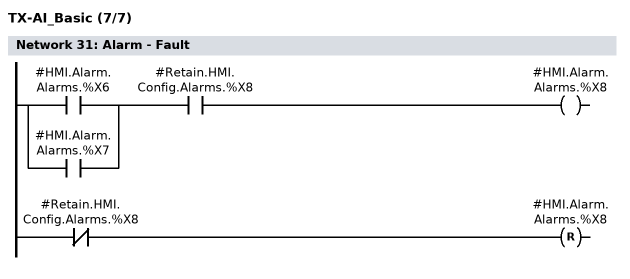
   RUNG wire#powerrail
      Contact( #HMI.Alarm.Alarms.%X6 )
      wire#w1
      Contact( #Retain.HMI.Config.Alarms.%X8 )
      Coil( #HMI.Alarm.Alarms.%X8 )
   END_RUNG
   RUNG wire#powerrail
      Contact( #HMI.Alarm.Alarms.%X7 )
   END_RUNG wire#w1
   RUNG wire#powerrail
      I_Contact( #Retain.HMI.Config.Alarms.%X8 )
      R_Coil( #HMI.Alarm.Alarms.%X8 )
   END_RUNG
   // the same network as SCL:
   #HMI.Alarm.Alarms.%X8 := (#HMI.Alarm.Alarms.%X6 OR #HMI.Alarm.Alarms.%X7) AND #Retain.HMI.Config.Alarms.%X8;
   IF NOT #Retain.HMI.Config.Alarms.%X8 THEN #HMI.Alarm.Alarms.%X8 := FALSE; END_IF;
END_REGION

REGION Network 32 (SCL)
   #Alarms.HighHighHigh := #HMI.Alarm.Alarms.%X0;
   #Alarms.HighHigh := #HMI.Alarm.Alarms.%X1;
   #Alarms.High := #HMI.Alarm.Alarms.%X2;
   #Alarms.Low := #HMI.Alarm.Alarms.%X3;
   #Alarms.LowLow := #HMI.Alarm.Alarms.%X4;
   #Alarms.LowLowLow := #HMI.Alarm.Alarms.%X5;
   #Alarms.OverRange := #HMI.Alarm.Alarms.%X6;
   #Alarms.UnderRange := #HMI.Alarm.Alarms.%X7;
   #Alarms.TransmitterFault := #HMI.Alarm.Alarms.%X8;
END_REGION
END_FUNCTION_BLOCK

FUNCTION_BLOCK "2oo3 AI"   // FB880, LAD
{ S7_Optimized_Access := 'TRUE' }
VERSION : 0.1
   VAR_INPUT
      V1GA : Bool;   // Value 1
      V2GA : Bool;   // Value 2
      V3GA : Bool;   // Value 3
      "2oo3.HH" : Bool;
      "2oo3.H" : Bool;
      "2oo3.L" : Bool;
      "2oo3.LL" : Bool;
      "2oo3.Trip" : Bool;
      PM : Int;   // Permissive Mode - "0=No P""1=Bool P" "2=Real P"
      HPB : Bool := TRUE;   // High Permissive BOOL
      LPB : Bool := TRUE;   // Low Permissive BOOL
      HPR : Real;   // High Permissive REAL
      LPR : Real;   // Low Permissive REAL
   END_VAR
   VAR_OUTPUT
      V1GA_1 : Bool;   // Value 1
      V2GA_1 : Bool;   // Value 2
      V3GA_1 : Bool;   // Value 3
      "2oo3.HH_1" : Bool;
      "2oo3.H_1" : Bool;
      "2oo3.L_1" : Bool;
      "2oo3.Trip_1" : Bool;
      "2oo3.LL_1" : Bool;
   END_VAR
   VAR
      Config : Struct   // Configurations
         Limits : Struct
            HH : Real := 100.0;   // High High Limit
            H : Real := 90.0;   // High Limit
            L : Real := 10.0;   // Low Limit
            LL : Real := 5.0;   // Low Low Limit
         END_STRUCT;
         H : Real := 1.0;   // Hysteresis
      END_STRUCT;
      Alarms : Struct
         HH : Bool;   // High High
         H : Bool;   // High
         L : Bool;   // Low
         LL : Bool;   // Low Low
         V1GA : Bool;   // Value 1 General Alarm
         V2GA : Bool;   // Value 2 General Alarm
         V3GA : Bool;   // Value 3 General Alarm
      END_STRUCT;
      "HMI.FVR" : Real := 100.0;
      "FVR.HH" : DInt;
      "FVR.H" : DInt;
      "FVR.L" : DInt;
      "FVR.LL" : DInt;
      "FVR.HPR" : DInt;
      "FVR.LPR" : DInt;
      "FVR.CONFIG.H" : DInt;
   END_VAR
   VAR_TEMP
      "MATH.HH" : Real;
      "MATH.H" : Real;
      "MATH.LL" : Real;
      "MATH.L" : Real;
      "MATH.HR" : Real;
      "MATH.LR" : Real;
      "MATH.CONFIG.H" : Real;
   END_VAR
BEGIN

REGION Network 1
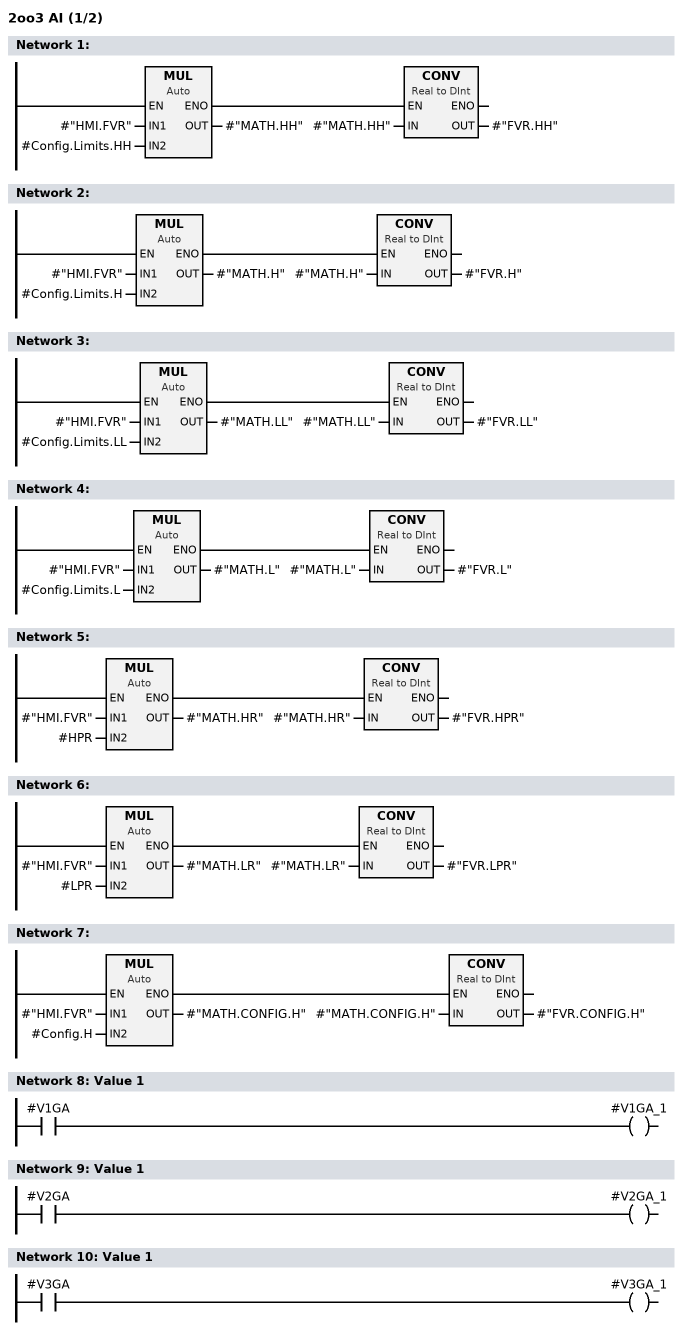
   RUNG wire#powerrail
      Mul(in1 := #"HMI.FVR", in2 := #Config.Limits.HH, out => #"MATH.HH")
      { S7_Templates := "[SrcType := Real, DestType := DInt]" } Convert(in := #"MATH.HH", out => #"FVR.HH")
   END_RUNG
   // the same network as SCL:
   #"MATH.HH" := #"HMI.FVR" * #Config.Limits.HH;
   #"FVR.HH" := REAL_TO_DINT(#"MATH.HH");
END_REGION

REGION Network 2
   RUNG wire#powerrail
      Mul(in1 := #"HMI.FVR", in2 := #Config.Limits.H, out => #"MATH.H")
      { S7_Templates := "[SrcType := Real, DestType := DInt]" } Convert(in := #"MATH.H", out => #"FVR.H")
   END_RUNG
   // the same network as SCL:
   #"MATH.H" := #"HMI.FVR" * #Config.Limits.H;
   #"FVR.H" := REAL_TO_DINT(#"MATH.H");
END_REGION
